(* Logix 5000 project; controller PLC_MCC1300_75F1 vendor 1 type 14 code 166 rev 32.11; software revision 32.04 *)

TASK _18_STI (periodic, rate 10 ms, priority 10, watchdog 500 ms) : _18_STI
TASK Diagnostic (periodic, rate 500 ms, priority 15, watchdog 2000 ms) : Modules
TASK MainTask (periodic, rate 6 ms, priority 10, watchdog 500 ms) : Initialize, MainProgram, CommandLogic, MotionLogic, Communication

MODULES
   Local : vendor 1 type 14 code 166 (ICP 0, rev 32.11)
      ETH_MCC1300 : 1756-EN2T (ICP 1, Ethernet 138.84.12.118, rev 11.1)
         ETH_M2 : 1756-EN2T (Ethernet 138.84.12.123, rev 10.7)   // Plant Network
             : 1756-IB16 (ICP 2, rev 3.4, Input RPI 20 ms)
             : 1756-IB16 (ICP 6, rev 3.4, Input RPI 20 ms)
             : 1756-IB16 (ICP 3, rev 3.4, Input RPI 20 ms)
             : 1756-IB16 (ICP 4, rev 3.4, Input RPI 20 ms)
             : 1756-IB16 (ICP 5, rev 3.4, Input RPI 20 ms)
             : vendor 1 type 7 code 16 (ICP 11, rev 3.4, Output RPI 20 ms)
                 ETH_M2:11:O.Data   // Local output updates
            Rio_Loops_2_3 : 1756-DHRIO (ICP 13, rev 7.2, Input RPI 25 ms)
               VMCC_TD : 1771-ASB (RIO 8, rev 1.1, Output RPI 48 ms)
                    VMCC_TD:O   // RACK 2 OUTPUT UPDATES
               VMCC_M2CM01_SPEED : vendor 1 type 12 code 51 (RIO 13, rev 1.1, Output RPI 48 ms)
                    VMCC_M2CM01_SPEED:O   // RACK 3 OUPUT UPDATES
               VMCC_M2_M2CM02_Speed : vendor 1 type 12 code 51 (RIO 14, rev 1.1, Output RPI 48 ms)
                    VMCC_M2_M2CM02_Speed:O   // RACK 3 OUPUT UPDATES
               ROCKWELL_CAPPING_SYSTEM : vendor 1 type 12 code 51 (RIO 12, rev 1.1, Output RPI 48 ms)
                    ROCKWELL_CAPPING_SYSTEM:O   // RACK 3 OUPUT UPDATES
               PANEL_KD_CS1N : vendor 1 type 12 code 51 (RIO 16, rev 1.1, Output RPI 48 ms)
                    PANEL_KD_CS1N:O   // RACK 11 OUPUT UPDATES
               VMCC_M2_M2CM03_Speed : vendor 1 type 12 code 51 (RIO 15, rev 1.1, Output RPI 48 ms)
                    VMCC_M2_M2CM03_Speed:O   // RACK 3 OUPUT UPDATES
               PANEL_TD_CS1N : 1794-ASB (RIO 18, rev 1.1, Output RPI 48 ms)   // Trim knocker 1
                    PANEL_TD_CS1N:O   // RACK 4 OUPUT UPDATES
               Panel_TS_CS2N : vendor 1 type 12 code 51 (RIO 20, rev 1.1, Output RPI 48 ms)
                    Panel_TS_CS2N:O   // RACK 5 OUPUT UPDATES
               PANEL_TD_CS3N : vendor 1 type 12 code 51 (RIO 22, rev 1.1, Output RPI 48 ms)
                    PANEL_TD_CS3N:O   // RACK 5 OUPUT UPDATES
               PANEL_TD_CS4N : vendor 1 type 12 code 51 (RIO 24, rev 1.1, Output RPI 48 ms)
                    PANEL_TD_CS4N:O   // RACK 6 OUPUT UPDATES
               PANEL_TD_CS5N : vendor 1 type 12 code 51 (RIO 26, rev 1.1, Output RPI 48 ms)
                    PANEL_TD_CS5N:O   // RACK 6 OUPUT UPDATES
               PANEL_TD_CS5S : vendor 1 type 12 code 51 (RIO 28, rev 1.1, Output RPI 48 ms)
                    PANEL_TD_CS5S:I.Data[0].15   // Panel-TD-CS5S Relicance Handoff Sensor (Redundant Sensor on South Side)
                    PANEL_TD_CS5S:O   // RACK 7 OUPUT UPDATES
               PANEL_TD_CS4S : vendor 1 type 12 code 51 (RIO 30, rev 1.1, Output RPI 48 ms)
                    PANEL_TD_CS4S:O   // RACK 7 OUPUT UPDATES
               PANEL_TD_CS3S : vendor 1 type 12 code 51 (RIO 32, rev 1.1, Output RPI 48 ms)
                    PANEL_TD_CS3S:O   // RACK 10 OUPUT UPDATES
               PANEL_TD_CS2S : vendor 1 type 12 code 51 (RIO 34, rev 1.1, Output RPI 48 ms)
                    PANEL_TD_CS2S:O   // RACK 10 OUPUT UPDATES
               BENCHBOARD : vendor 1 type 12 code 51 (RIO 36, rev 1.1, Output RPI 48 ms)
                    BENCHBOARD:O   // RACK 11 OUPUT UPDATES
               PANEL_KD_CS1S : vendor 1 type 12 code 51 (RIO 38, rev 1.1, Output RPI 48 ms)
               PANEL_TD_CS1S : vendor 1 type 12 code 51 (RIO 40, rev 1.1, Output RPI 48 ms)
                    PANEL_TD_CS1S:O   // RACK 12 OUPUT UPDATES
               VMCC_M2CM4S : vendor 1 type 12 code 51 (RIO 42, rev 1.1, Output RPI 48 ms)
                    VMCC_M2CM4S:O   // RACK 12 OUPUT UPDATES
               VMCC_M2_M2CM4N : vendor 1 type 12 code 51 (RIO 43, rev 1.1, Output RPI 48 ms)
                    VMCC_M2_M2CM4N:O   // RACK 12 OUPUT UPDATES
               VMCC_M2_M2CM9S : vendor 1 type 12 code 51 (RIO 52, rev 1.1, Output RPI 48 ms)
                    VMCC_M2_M2CM9S:O   // RACK 15 OUPUT UPDATES
               VMCC_M2_M2CM9N : vendor 1 type 12 code 51 (RIO 53, rev 1.1, Output RPI 48 ms)
                    VMCC_M2_M2CM9N:O   // RACK 15 OUPUT UPDATES
               VMCC_M2_M2CM10S : vendor 1 type 12 code 51 (RIO 54, rev 1.1, Output RPI 48 ms)
                    VMCC_M2_M2CM10S:O   // RACK 15 OUPUT UPDATES
               VMCC_M2_M2CM10N : vendor 1 type 12 code 51 (RIO 55, rev 1.1, Output RPI 48 ms)
                    VMCC_M2_M2CM10N:O   // RACK 15 OUPUT UPDATES
               VMCC_M2_M2CM11S : vendor 1 type 12 code 51 (RIO 56, rev 1.1, Output RPI 48 ms)
                    VMCC_M2_M2CM11S:O   // RACK 16 OUPUT UPDATES
               VMCC_M2_M2CM11N : vendor 1 type 12 code 51 (RIO 57, rev 1.1, Output RPI 48 ms)
                    VMCC_M2_M2CM11N:O   // RACK 16 OUPUT UPDATES
               VMCC_M2_M2CM12S : vendor 1 type 12 code 51 (RIO 58, rev 1.1, Output RPI 48 ms)
                    VMCC_M2_M2CM12S:O   // RACK 16 OUPUT UPDATES
               VMCC_M2_M2CM12N : vendor 1 type 12 code 51 (RIO 59, rev 1.1, Output RPI 48 ms)
                    VMCC_M2_M2CM12N:O   // RACK 16 OUPUT UPDATES
               MB : vendor 1 type 12 code 51 (RIO 60, rev 1.1, Output RPI 48 ms)
                    MB:O   // RACK 17 OUPUT UPDATES
               VMCC_M2_M2CM5S : vendor 1 type 12 code 51 (RIO 44, rev 1.1, Output RPI 48 ms)
                    VMCC_M2_M2CM5S:O   // RACK 13 OUPUT UPDATES
               VMCC_M2_M2CM5N : vendor 1 type 12 code 51 (RIO 45, rev 1.1, Output RPI 48 ms)
                    VMCC_M2_M2CM5N:O   // RACK 13 OUPUT UPDATES
               VMCC_M2_M2CM6S : vendor 1 type 12 code 51 (RIO 46, rev 1.1, Output RPI 48 ms)
                    VMCC_M2_M2CM6S:O   // RACK 13 OUPUT UPDATES
               VMCC_M2_M2CM6N : vendor 1 type 12 code 51 (RIO 47, rev 1.1, Output RPI 48 ms)
                    VMCC_M2_M2CM6N:O   // RACK 13 OUPUT UPDATES
               VMCC_M2_M2CM7S : vendor 1 type 12 code 51 (RIO 48, rev 1.1, Output RPI 48 ms)
                    VMCC_M2_M2CM7S:O   // RACK 14 OUPUT UPDATES
               VMCC_M2_M2CM7N : vendor 1 type 12 code 51 (RIO 49, rev 1.1, Output RPI 48 ms)
                    VMCC_M2_M2CM7N:O   // RACK 14 OUPUT UPDATES
               VMCC_M2_M2CM8S : vendor 1 type 12 code 51 (RIO 50, rev 1.1, Output RPI 48 ms)
                    VMCC_M2_M2CM8S:O   // RACK 14 OUPUT UPDATES
               VMCC_M2_M2CM8N : vendor 1 type 12 code 51 (RIO 51, rev 1.1, Output RPI 48 ms)
                    VMCC_M2_M2CM8N:O   // RACK 14 OUPUT UPDATES
      RIOM13 : 1794-AENTR (Ethernet 192.168.36.11, rev 1.1, Output RPI 20 ms)
         R03_S00 : 1794-IB16 (Flex 0, rev 1.1)
         R03_S01 : 1794-IB16 (Flex 1, rev 1.1)
         R03_S02 : vendor 1 type 7 code 35 (Flex 2, rev 1.1)
      E73AZ1 : vendor 1 type 37 code 49 (Ethernet 192.168.32.131, rev 7.1, MotionDiagnostics RPI 1 ms, MotionSync RPI 1 ms)
      E93AZ1 : vendor 1 type 37 code 49 (Ethernet 192.168.32.132, rev 7.1, MotionDiagnostics RPI 1 ms)
      E53AZ1 : vendor 1 type 45 code 15 (Ethernet 192.168.32.101, rev 2.3, AMotionDiagnostics RPI 1 ms)
      E61AZ1 : vendor 1 type 45 code 15 (Ethernet 192.168.32.102, rev 2.3, AMotionDiagnostics RPI 1 ms)
      E62AZ1 : vendor 1 type 45 code 15 (Ethernet 192.168.32.103, rev 2.3, AMotionDiagnostics RPI 1 ms)
      E63AZ1 : vendor 1 type 45 code 15 (Ethernet 192.168.32.104, rev 2.3, AMotionDiagnostics RPI 1 ms)
      E64AZ1 : vendor 1 type 45 code 15 (Ethernet 192.168.32.105, rev 2.3, AMotionDiagnostics RPI 1 ms)
      E65AZ1 : vendor 1 type 45 code 15 (Ethernet 192.168.32.106, rev 2.3, AMotionDiagnostics RPI 1 ms)
      E66AZ1 : vendor 1 type 45 code 15 (Ethernet 192.168.32.107, rev 2.3, AMotionDiagnostics RPI 1 ms)
      E67AZ1 : vendor 1 type 45 code 15 (Ethernet 192.168.32.108, rev 2.3, AMotionDiagnostics RPI 1 ms)
      E71AZ1 : vendor 1 type 45 code 15 (Ethernet 192.168.32.109, rev 2.3, AMotionDiagnostics RPI 1 ms)
      E76AZ1 : vendor 1 type 45 code 15 (Ethernet 192.168.32.110, rev 2.3, AMotionDiagnostics RPI 1 ms)
      E77AZ1 : vendor 1 type 45 code 15 (Ethernet 192.168.32.111, rev 2.3, AMotionDiagnostics RPI 1 ms)
      E78AZ1 : vendor 1 type 45 code 15 (Ethernet 192.168.32.112, rev 2.3, AMotionDiagnostics RPI 1 ms)
      E81AZ1 : vendor 1 type 45 code 15 (Ethernet 192.168.32.113, rev 2.3, AMotionDiagnostics RPI 1 ms)
      E82AZ1 : vendor 1 type 45 code 15 (Ethernet 192.168.32.114, rev 2.3, AMotionDiagnostics RPI 1 ms)
      E83AZ1 : vendor 1 type 45 code 15 (Ethernet 192.168.32.115, rev 2.3, AMotionDiagnostics RPI 1 ms)
      E84AZ1 : vendor 1 type 45 code 15 (Ethernet 192.168.32.116, rev 2.3, AMotionDiagnostics RPI 1 ms)
      E85AZ1 : vendor 1 type 45 code 15 (Ethernet 192.168.32.117, rev 2.3, AMotionDiagnostics RPI 1 ms)
      E86AZ1 : vendor 1 type 45 code 15 (Ethernet 192.168.32.118, rev 2.3, AMotionDiagnostics RPI 1 ms)
      E87AZ1 : vendor 1 type 45 code 15 (Ethernet 192.168.32.119, rev 2.3, AMotionDiagnostics RPI 1 ms)
      E88AZ1 : vendor 1 type 45 code 15 (Ethernet 192.168.32.120, rev 2.3, AMotionDiagnostics RPI 1 ms)
      E91AZ1 : vendor 1 type 45 code 15 (Ethernet 192.168.32.121, rev 2.3, AMotionDiagnostics RPI 1 ms)
      E96AZ1 : vendor 1 type 45 code 15 (Ethernet 192.168.32.122, rev 2.3, AMotionDiagnostics RPI 1 ms)
      E97AZ1 : vendor 1 type 45 code 15 (Ethernet 192.168.32.123, rev 2.3, AMotionDiagnostics RPI 1 ms)
      E98AZ1 : vendor 1 type 45 code 15 (Ethernet 192.168.32.124, rev 2.3, AMotionDiagnostics RPI 1 ms)
      M3AZ01 : vendor 1 type 45 code 15 (Ethernet 192.168.32.141, rev 2.3, AMotionDiagnostics RPI 1 ms)
      M3AZ02 : vendor 1 type 45 code 15 (Ethernet 192.168.32.142, rev 2.3, AMotionDiagnostics RPI 1 ms)
      M3AZ03 : vendor 1 type 45 code 15 (Ethernet 192.168.32.143, rev 2.3, AMotionDiagnostics RPI 1 ms)
      M3AZ04 : vendor 1 type 45 code 15 (Ethernet 192.168.32.144, rev 2.3, AMotionDiagnostics RPI 1 ms)
      M3AZ05 : vendor 1 type 45 code 15 (Ethernet 192.168.32.145, rev 2.3, AMotionDiagnostics RPI 1 ms)
      M3AZ06 : vendor 1 type 45 code 15 (Ethernet 192.168.32.146, rev 2.3, AMotionDiagnostics RPI 1 ms)
      M3AZ07 : vendor 1 type 45 code 15 (Ethernet 192.168.32.147, rev 2.3, AMotionDiagnostics RPI 1 ms)
      M3AZ08 : vendor 1 type 45 code 15 (Ethernet 192.168.32.148, rev 2.3, AMotionDiagnostics RPI 1 ms)
      M3AZ09 : vendor 1 type 45 code 15 (Ethernet 192.168.32.149, rev 2.3, AMotionDiagnostics RPI 1 ms)
      M3AZ10 : vendor 1 type 45 code 15 (Ethernet 192.168.32.150, rev 2.3, AMotionDiagnostics RPI 1 ms)
      D010M1PM1 : vendor 1 type 45 code 15 (Ethernet 192.168.36.131, rev 2.3, AMotionDiagnostics RPI 1 ms)
      D010M2PM1 : vendor 1 type 45 code 15 (Ethernet 192.168.36.132, rev 2.3, AMotionDiagnostics RPI 1 ms)
      D020M1PM1 : vendor 1 type 45 code 15 (Ethernet 192.168.36.133, rev 2.3, AMotionDiagnostics RPI 1 ms)
      TDKAZ00N : vendor 1 type 45 code 15 (Ethernet 192.168.31.101, rev 2.3, AMotionDiagnostics RPI 1 ms)
      TDKAZ00S : vendor 1 type 45 code 15 (Ethernet 192.168.31.102, rev 2.3, AMotionDiagnostics RPI 1 ms)
      TDKAZ01N : vendor 1 type 45 code 15 (Ethernet 192.168.31.103, rev 2.3, AMotionDiagnostics RPI 1 ms)
      TDKAZ01S : vendor 1 type 45 code 15 (Ethernet 192.168.31.104, rev 2.3, AMotionDiagnostics RPI 1 ms)
      TDKAZ02N : vendor 1 type 45 code 15 (Ethernet 192.168.31.105, rev 2.3, AMotionDiagnostics RPI 1 ms)
      TDKAZ02S : vendor 1 type 45 code 15 (Ethernet 192.168.31.106, rev 2.3, AMotionDiagnostics RPI 1 ms)
      TDKAZ03N : vendor 1 type 45 code 15 (Ethernet 192.168.31.107, rev 2.3, AMotionDiagnostics RPI 1 ms)
      TDKAZ03S : vendor 1 type 45 code 15 (Ethernet 192.168.31.108, rev 2.3, AMotionDiagnostics RPI 1 ms)
      TDKAZ04N : vendor 1 type 45 code 15 (Ethernet 192.168.31.109, rev 2.3, AMotionDiagnostics RPI 1 ms)
      TDKAZ04S : vendor 1 type 45 code 15 (Ethernet 192.168.31.110, rev 2.3, AMotionDiagnostics RPI 1 ms)
      TDKAZ05N : vendor 1 type 45 code 15 (Ethernet 192.168.31.111, rev 2.3, AMotionDiagnostics RPI 1 ms)
      TDKAZ05S : vendor 1 type 45 code 15 (Ethernet 192.168.31.112, rev 2.3, AMotionDiagnostics RPI 1 ms)
      TDAZ00N : vendor 1 type 45 code 15 (Ethernet 192.168.31.113, rev 2.3, AMotionDiagnostics RPI 1 ms)
      TDAZ00S : vendor 1 type 45 code 15 (Ethernet 192.168.31.114, rev 2.3, AMotionDiagnostics RPI 1 ms)
      TDAZ01N : vendor 1 type 45 code 15 (Ethernet 192.168.31.115, rev 2.3, AMotionDiagnostics RPI 1 ms)
      TDAZ01S : vendor 1 type 45 code 15 (Ethernet 192.168.31.116, rev 2.3, AMotionDiagnostics RPI 1 ms)
      TDAZ02N : vendor 1 type 45 code 15 (Ethernet 192.168.31.117, rev 2.3, AMotionDiagnostics RPI 1 ms)
      TDAZ02S : vendor 1 type 45 code 15 (Ethernet 192.168.31.118, rev 2.3, AMotionDiagnostics RPI 1 ms)
      TDAZ03N : vendor 1 type 45 code 15 (Ethernet 192.168.31.119, rev 2.3, AMotionDiagnostics RPI 1 ms)
      TDAZ03S : vendor 1 type 45 code 15 (Ethernet 192.168.31.120, rev 2.3, AMotionDiagnostics RPI 1 ms)
      TDAZ04N : vendor 1 type 45 code 15 (Ethernet 192.168.31.121, rev 2.3, AMotionDiagnostics RPI 1 ms)
      TDAZ04S : vendor 1 type 45 code 15 (Ethernet 192.168.31.122, rev 2.3, AMotionDiagnostics RPI 1 ms)
      TDAZ05N : vendor 1 type 45 code 15 (Ethernet 192.168.31.123, rev 2.3, AMotionDiagnostics RPI 1 ms)
      TDAZ05S : vendor 1 type 45 code 15 (Ethernet 192.168.31.124, rev 2.3, AMotionDiagnostics RPI 1 ms)
      E152AP1 : vendor 1 type 12 code 317 (Ethernet 192.168.32.11, rev 4.1)
         R00_S03 : 5069-IB16 (5069 3, rev 2.1, StandardDataDriven RPI 5 ms)
         R00_S04 : 5069-IB16 (5069 4, rev 2.1, StandardDataDriven RPI 5 ms)
         R00_S02 : 5069-IB16 (5069 2, rev 2.1, StandardDataDriven RPI 5 ms)
         R00_S01 : 5069-IB16 (5069 1, rev 2.1, StandardDataDriven RPI 5 ms)
         R00_S05 : 5069-IB16 (5069 5, rev 2.1, StandardDataDriven RPI 5 ms)
         R00_S06 : 5069-IB16 (5069 6, rev 2.1, StandardDataDriven RPI 5 ms)
         R00_S07 : 5069-IB16 (5069 7, rev 2.1, StandardDataDriven RPI 5 ms)
         R00_S08 : 5069-IB16 (5069 8, rev 2.1, StandardDataDriven RPI 5 ms)
         R00_S09 : 5069-IB16 (5069 9, rev 2.1, StandardDataDriven RPI 5 ms)
         R00_S10 : 5069-IB16 (5069 10, rev 2.1, StandardDataDriven RPI 5 ms)
         R00_S11 : 5069-IB16 (5069 11, rev 2.1, StandardDataDriven RPI 5 ms)
         R00_S12 : 5069-IB16 (5069 12, rev 2.1, StandardDataDriven RPI 5 ms)
         R00_S13 : 5069-OB16 (5069 13, rev 3.1, StandardDataDriven RPI 5 ms)
         R00_S14 : 5069-OB16 (5069 14, rev 3.1, StandardDataDriven RPI 5 ms)
         R00_S15 : 5069-OB16 (5069 15, rev 3.1, StandardDataDriven RPI 5 ms)
         R00_S16 : 5069-OB16 (5069 16, rev 3.1, StandardDataDriven RPI 5 ms)
         R00_S17 : 5069-OB16 (5069 17, rev 3.1, StandardDataDriven RPI 5 ms)
      M3683AP1 : vendor 1 type 12 code 317 (Ethernet 192.168.31.12, rev 4.1)
         R01_S01 : 5069-IB16 (5069 1, rev 2.1, StandardDataDriven RPI 5 ms)
         R01_S02 : 5069-IB16 (5069 2, rev 2.1, StandardDataDriven RPI 5 ms)
         R01_S03 : 5069-IB16 (5069 3, rev 2.1, StandardDataDriven RPI 5 ms)
         R01_S04 : 5069-IB16 (5069 4, rev 2.1, StandardDataDriven RPI 5 ms)
         R01_S05 : 5069-OB16 (5069 5, rev 3.1, StandardDataDriven RPI 5 ms)
         R01_S06 : 5069-OB16 (5069 6, rev 3.1, StandardDataDriven RPI 5 ms)
         R01_S07 : 5069-OB16 (5069 7, rev 3.1, StandardDataDriven RPI 5 ms)
         R01_S08 : 5069-OB16 (5069 8, rev 3.1, StandardDataDriven RPI 5 ms)
         R01_S09 : 5069-OB16 (5069 9, rev 3.1, StandardDataDriven RPI 5 ms)
         R01_S10 : 5069-IB16 (5069 10, rev 2.1, StandardDataDriven RPI 5 ms)
      TD5680AP1 : vendor 1 type 12 code 317 (Ethernet 192.168.31.11, rev 4.1)
         R02_S01 : 5069-IB16 (5069 1, rev 2.1, StandardDataDriven RPI 5 ms)
         R02_S02 : 5069-IB16 (5069 2, rev 2.1, StandardDataDriven RPI 5 ms)
         R02_S03 : 5069-OB16 (5069 3, rev 3.1, StandardDataDriven RPI 5 ms)
         R02_S04 : 5069-OB16 (5069 4, rev 3.1, StandardDataDriven RPI 5 ms)
         R02_S05 : 5069-OB16 (5069 5, rev 3.1, StandardDataDriven RPI 5 ms)
         R02_S06 : 5069-OB16 (5069 6, rev 3.1, StandardDataDriven RPI 5 ms)
         R02_S07 : 5069-IB16 (5069 7, rev 2.1, StandardDataDriven RPI 5 ms)
         R02_S08 : 5069-IB16 (5069 8, rev 2.1, StandardDataDriven RPI 5 ms)
END_MODULES

TYPE AUX_COSTANTS :
STRUCT
   dM302SnapOffset_cmm : DINT;   // Distance from origin sepoint and snapbar [mm/100]
   dM302SpeedUpMinGapInConvoy_cmm : DINT;   // Minimum gap in convoy [mm/100]
   dM310_PopUpCycleTime_s : DINT[2];   // Popup cycle time [s]
   dM315_PopUpCycleTime_s : DINT[2];   // Popup cycle time [s]
END_STRUCT
END_TYPE

TYPE CM_AreaStackerToLine :
STRUCT
   dSyncHead : DINT;
   xRequestAccessArea : BOOL;
   xAccessAreaAccepted : BOOL;
   xAreaOk : BOOL;
   xStackerInUnloaderMode : BOOL;
   xStackerInProduction : BOOL;
   xPlateOnFrame : BOOL[32];
   xSB_SilenceAlarm : BOOL;
   xSB_SendToCullet : BOOL;
   xSB_LineCycle : BOOL;
   xSB_StopLineCycle : BOOL;
   xSB_LineJogPlus : BOOL;
   xSB_LineJogMinus : BOOL;
   xSB_DestinationChange : BOOL;
   iPresetNumberPlateOnRack : INT[2];
   iActualNumberPlateOnRack : INT[2];
   iPresetNumberPlateAddOnRack : INT[2];
   iActualNumberPlateAddOnRack : INT[2];
   dGap_cmm : DINT;
   dMsgDataSyncFdbk : DINT;
   dMsgDataSync : DINT;
   dMsgOPTSyncFdbk : DINT;
   dMsgOPTSync : DINT;
   dSyncTail : DINT;
END_STRUCT
END_TYPE

TYPE CM_ConveyorStackerToLine :
STRUCT
   dSyncHead : DINT;
   xCycleOn : BOOL;
   xConditionOkForStopCycle : BOOL;
   xInitialContionOk : BOOL;
   xOutputEnable : BOOL;
   xReadyToMove : BOOL;
   xFeedbackRotation : BOOL;
   xRequestReturnInLine : BOOL;
   xRequestUnload : BOOL;
   xRotationForUnload : BOOL;
   xRotationForLoad : BOOL;
   xEndPhaseLoad : BOOL;
   xManualCommandFwd : BOOL;
   xManualCommandBkw : BOOL;
   xAirMode : BOOL;
   xTinMode : BOOL;
   xPhotocell1 : BOOL;
   xPhotocell2 : BOOL;
   xPlateOnConveyor : BOOL[32];
   dSyncTail : DINT;
END_STRUCT
END_TYPE

TYPE CM_DATA_Z200 :   // Cap data coming from Z200
STRUCT
   dSyncHead : DINT;   // Synchro head
   tConvoyCap : UDT_ConvoyCap_ZC;   // Cap data
   dSyncTail : DINT;   // Synchro tail
END_STRUCT
END_TYPE

TYPE CM_INPUT_Z200 :
STRUCT
   dSyncHead : DINT;   // Synchro head
   xZ200_CycleON : BOOL;   // Z200 Cycle ON
   xSnapDone : BOOL;   // Snap done
   xSBStartEmptyingZ301 : BOOL;   // CS4201 Start Emptying Z301 Button
   xSBStopEmptyingZ301 : BOOL;   // CS4201 Stop Emptying Z301 Button
   xSBResetAnomalyZ301 : BOOL;   // CS4201 Reset Anomaly Z301 Button
   xResetGeneralEmergency : BOOL;   // Reset General Emergency
   xCrossbreakActive : BOOL;   // Crossbreak Active
   xEmergencyON : BOOL;   // Emergency ON
   xMainCulletConveyorAllow : BOOL;   // Main Cullet Conveyor Allow
   dLehrSpeed_mm_min : DINT;   // Lehr speed [mm/min]
   dDataSync : DINT;   // Snap cap data sent
   rgdSpare : DINT[10];
   dSyncTail : DINT;   // Synchro tail
END_STRUCT
END_TYPE

TYPE CM_LineToAreaStacker :
STRUCT
   dSyncHead : DINT;
   xConditionOkForAccessArea : BOOL;
   xSBSendToCullet : BOOL;
   xSBLineCycle : BOOL;
   xSBStopLineCycle : BOOL;
   xHLAlarmStartLineCycle : BOOL;
   xSBChangeDestination : BOOL;
   dMsgDataSyncFdbk : DINT;
   dMsgDataSync : DINT;
   dMsgOPTSyncFdbk : DINT;
   dMsgOPTSync : DINT;
   dSyncTail : DINT;
END_STRUCT
END_TYPE

TYPE CM_LineToConveyorStacker :
STRUCT
   dSyncHead : DINT;
   xEmergencyOn : BOOL;
   xLineCycleOn : BOOL;
   xLineStopCycle : BOOL;
   xRequestForceStop : BOOL;
   xResetAlarms : BOOL;
   xResetEmergency : BOOL;
   xPowerOnByLine : BOOL;
   xInitialConditionOk : BOOL;
   xOutputEnable : BOOL;
   xReadyToMove : BOOL;
   xFeedbackRotation : BOOL;
   xEndPhaseLoad : BOOL;
   xRotationForLoad : BOOL;
   xRequestForUnload : BOOL;
   xRotationForUnload : BOOL;
   xManualCommandFwd : BOOL;
   xManualCommandBkw : BOOL;
   xSendToCullet : BOOL;
   xLineJogPlus : BOOL;
   xLineJogMinus : BOOL;
   dLineSpeed_dmm_min : DINT;
   dSyncTail : DINT;
END_STRUCT
END_TYPE

TYPE CM_OUTPUT_Z200 :
STRUCT
   dSyncHead : DINT;   // Synchro head
   xZ300_CycleON : BOOL;   // Z300 Cycle ON
   xBLStartEmptyingZ301Light : BOOL;   // CS4201 Start Emptying Z301 Button Light
   xBLStopEmptyingZ301Light : BOOL;   // CS4201 Stop Emptying Z301 Button Light
   xBLAnomalyZ301Light : BOOL;   // CS4201 Anomaly Z301 Button Light
   xBLAnomalyZ302Light : BOOL;   // CS4201 Anomaly Z302 Button Light
   dDataSyncFdbk : DINT;   // Snap cap sync feedback
   dLineSpeed_mm_min : DINT;   // Line speed [mm/min]
   rgdSpare : DINT[10];
   dSyncTail : DINT;   // Synchro tail
END_STRUCT
END_TYPE

TYPE DATA_CAP_PILKINGTON :
STRUCT
   dHost_ID : DINT;   // Host ID
   dCap_Length_64ths : DINT;   // Cap Length (64ths)
   dCap_Primary_Destination_Mask : DINT;   // Cap Primary Destination Mask
   Packing_station_1_Mask : DINT;   // Packing Station 1 Mask
   Packing_station_2_Mask : DINT;   // Packing Station 2 Mask
   Packing_station_3_Mask : DINT;   // Packing Station 3 Mask
   Packing_station_4_Mask : DINT;   // Packing Station 4 Mask
   Packing_station_5_Mask : DINT;   // Packing Station 5 Mask
   dSplit_A_Width_64ths : DINT;   // Split A Width (64ths)
   dSplit_A_Dest_Mask : DINT;   // Split A Destination Mask
   dSplit_B_Width_64ths : DINT;   // Split B Width (64ths)
   dSplit_B_Dest_Mask : DINT;   // Split B Destination Mask
   dSplit_C_Width_64ths : DINT;   // Split C Width (64ths)
   dSplit_C_Dest_Mask : DINT;   // Split C Destination Mask
   dSplit_D_Width_64ths : DINT;   // Split D Width (64ths)
   dSplit_D_Dest_Mask : DINT;   // Split D Destination Mask
   dCap_Secondary_Dest_Mask : DINT;   // Cap Secondary Destination Mask
   dTrim_Home_Side_64ths : DINT;   // Trim on home (left) side (64ths)
   dTrim_Far_Side_64ths : DINT;   // Trim on far (right) side (64ths)
   dControl_Bits_For_Legs : DINT;   // Control bits for legs
   dCap_Width_64ths : DINT;   // Cap Width (64ths)
   dReject_Mask : DINT;   // Split Reject mask
   dPattern_number : DINT;   // Pattern number
   dSpare1 : DINT;   // Spare
   dSpare2 : DINT;   // Spare
   dSpare3 : DINT;   // Spare
   dMainline_History_Word : DINT;   // Mainline History Word
   dSpare4 : DINT;   // Spare
   dSpare5 : DINT;   // Spare
   dSpare6 : DINT;   // Spare
   dSpare7 : DINT;   // Spare
   dSpare8 : DINT;   // Spare
   dSpare9 : DINT;   // Spare
END_STRUCT
END_TYPE

TYPE GP_AccessArea_STC :
STRUCT
   ST_xAccessRequest : BOOL;
   ST_xAccessAccepted : BOOL;
   ST_xAccessAnnulled : BOOL;
   ST_xAccessAcceptedAndButtonReleased : BOOL;
   ST_xConditionOkForAccess : BOOL;
   ST_xDelayForceAccess : BOOL;
   ST_xSafetyOkForCycle : BOOL;
   OSR_xAccessRequest : BOOL;
   OSR_xAccessAcceptedAndButtonReleased : BOOL;
   OSR_xRemoveAccess : BOOL;
   OSR_xRemoveAccessNotAccepted : BOOL;
   OS_xAccessRequest : BOOL;
   OS_xSafetyOK : BOOL;
   tmON_ForceAccess : TIMER;
END_STRUCT
END_TYPE

TYPE GP_NetworkDiag_v1 :
STRUCT
   sModuleName : STRING;   // Module name
   xConnected : BOOL;   // Module connected
   xFaulted : BOOL;   // Module faulted
   dEntryStatus : DINT;
   dFaultCode : DINT;
   dFaultInfo : DINT;
   dInstance : DINT;
END_STRUCT
END_TYPE

TYPE GP_OB_Initialize_STC :
STRUCT
   dElapsed_1h_ms : DINT;   // Decimal
   dElapsed_1min_ms : DINT;   // Decimal
   dElapsed_1s_ms : DINT;   // Decimal
   dElapsed_2min_ms : DINT;   // Decimal
   dElapsed_2s_ms : DINT;   // Decimal
   dElapsed_5s_ms : DINT;   // Decimal
   dElapsed_10min_ms : DINT;   // Decimal
   dElapsed_10s_ms : DINT;   // Decimal
   dElapsed_30min_ms : DINT;   // Decimal
   dElapsed_30s_ms : DINT;   // Decimal
   dElapsed_100ms_ms : DINT;   // Decimal
   dElapsed_200ms_ms : DINT;   // Decimal
   dElapsed_400ms_ms : DINT;   // Decimal
   dElapsed_500ms_ms : DINT;   // Decimal
   dElapsed_800ms_ms : DINT;   // Decimal
   dlLastExecValue_us : DINT;   // Decimal
   rReminder_ms : REAL;   // Float
   lwOldStartTime : DINT[2];   // Old start time execution
   lwStartTime : DINT[2];   // Start time execution
END_STRUCT
END_TYPE

TYPE GP_TrackingSearchPlate_STC :
STRUCT
   rgdHeadPointer : DINT[5];   // Head pointer
   rgdTailPointer : DINT[5];   // Tail pointer
   rgdHead_cmm : DINT[5];   // Head position [cmm]
   rgdTail_cmm : DINT[5];   // Tail position [cmm]
   rgxHead : DINT;   // Head found
   rgxTail : DINT;   // Tail found
   xHeadPresence : BOOL;   // At least one head
   xTailPresence : BOOL;   // At least one tail
END_STRUCT
END_TYPE

TYPE HMI_LiteData :
STRUCT
   dHead_PosX_mm : DINT;   // Plate head position X [mm]
   dTail_PosX_mm : DINT;   // Plate tail position X [mm]
   dPlateLength_mm : DINT;   // Plate length [mm]
   dPositionY_mm : DINT;   // Plate position Y [mm]- Operator side
   dPlateWidth_mm : DINT;   // Plate widht [mm]
   dPlateId : DINT;   // Plate ID
   dProductionID : DINT;   // Production ID
   dSource : DINT;   // Plate source
   dDestination : DINT;   // Plate Main destination
   dAlternative : DINT;   // Plate Alternative destination
   dSecondDestination : DINT;   // Plate 2nd choice destination
END_STRUCT
END_TYPE

TYPE MAC_Conveyor :
STRUCT
   ST_xInitialConditionOK : BOOL;   // Initial condition OK
   ST_xInitialConditionOK_BW : BOOL;   // Initial condition OK backward
   ST_xCleaningConditionOK : BOOL;   // Cleaning condition OK
   ST_xCleaningAccepted : BOOL;   // Cleaning accepted
   ST_xReqCleaning : BOOL;   // Request cleaning
   ST_xPlatePresence : BOOL;   // Plate presence memory
   ST_xPhasesInProgress : BOOL;   // Phases in progress
   ST_xCycleLoadUnload : BOOL;   // Cycle load/unload simultaneously
   ST_xStopMachineFault : BOOL;   // Stopped machine fault
   ST_xStopNextCycleFault : BOOL;   // Stop next cycle fault
   ST_xConditionOKStopCycle : BOOL;   // Condition OK for stop cycle
   ST_xOutputEnable : BOOL;   // Output enable
   ST_xMachineAlarm : BOOL;   // Machine alarm
   ST_xMachineWarning : BOOL;   // Machine warning
   ST_xIdPlatePresence : BOOL;   // Id plate presence
   ST_xFeedbackRotation : BOOL;   // Feedback rotation
   ST_xRampInProgress : BOOL;   // Ramp in progress
   ST_xAccInProgress : BOOL;   // Acceleration in progress
   ST_xDecInProgress : BOOL;   // Deceleration in progress
   ST_xWaitStopNextMachine : BOOL;   // Wait stop next machine
   ST_xWaitMachineStop : BOOL;   // Wait machine stop
   ST_xWaitReadyToMove : BOOL;   // Wait ready to move
   ST_xEnableControlError : BOOL;   // Enable control error
   ST_xManualMode : BOOL;   // Manual mode enabled
   ST_xPlateSynchronized : BOOL;   // Plate synchronized
   ST_xVirtualDoorEnabled : BOOL;   // Virtual door enabled
   ST_xDisableLoadUnloadOnStop : BOOL;   // Temporary disable of load/unload continuosly after a bit wait machine stop
   ST_xPlatePassageUpstream_FW : BOOL;   // Plate in passage upstream
   ST_xPlatePassageUpstream_BKW : BOOL;   // Plate in passage upstream
   ST_xPlatePassageDownstream_FW : BOOL;   // Plate in passage downstream
   ST_xPlatePassageDownstream_BKW : BOOL;   // Plate in passage downstream
   ST_xAxleReadyToMoveDelayed : BOOL;   // Axle ready to move delayed (NU)
   ST_xSafetyMovement : BOOL;   // Safety Mouvement
   ST_xReqDescent : BOOL;   // popup conveyor
   ST_xPhaseError : BOOL;   // Phase error, send lites to cullet
   ST_xAux1 : BOOL;   // ST Aux 1
   ST_xAux2 : BOOL;   // ST Aux 2
   ST_xAux3 : BOOL;   // ST Aux 3
   ST_xAux4 : BOOL;   // ST Aux 4
   OSR_xUnload : BOOL;   // OSR Unload
   OSR_xSynchroPhotocellHead : BOOL;   // OSR Synchronization photocell head
   OSR_xSynchroPhotocellTail : BOOL;   // OSR Synchronization photocell tail
   OSR_xPosReq : BOOL;   // OSR Positioning request
   OS_xLoad_FW : BOOL;   // OS Load forward
   OS_xUnload_FW : BOOL;   // OS Unload forward
   OS_xLoad_BW : BOOL;   // OS Load backward
   OS_xUnload_BW : BOOL;   // OS Unload backward
   OS_xUnpack : BOOL;   // OS Unpack convoy
   OS_xSynchroPhotocellHead : BOOL;   // OS Synchronization photocell head
   OS_xSynchroPhotocellTail : BOOL;   // OS Synchronization photocell tail
   OS_xChangeSpeed : BOOL;   // OS Dynamic change speed
   PH_x : DINT;   // Phases
   INPUT_xSyncroPhotocell_1 : BOOL;   // Sincro photocell / start count #1
   INPUT_xSyncroPhotocell_2 : BOOL;   // Sincro photocell / start count #2
   INPUT_xSquaringPhotocell_1 : BOOL;   // Squaring photocell #1
   INPUT_xSquaringPhotocell_2 : BOOL;   // Squaring photocell #2
   INPUT_xSquaringPhotocell_3 : BOOL;   // Squaring photocell #3
   INPUT_xSquaringPhotocell_4 : BOOL;   // Squaring photocell #4
   INPUT_xHighPositionSquaring_1 : BOOL;   // High position squaring #1
   INPUT_xLowPositionSquaring_1 : BOOL;   // Low position squaring #1
   INPUT_xHighPositionSquaring_2 : BOOL;   // High position squaring #2
   INPUT_xLowPositionSquaring_2 : BOOL;   // Low position squaring #2
   INPUT_xHighPositionPopup_1 : BOOL;   // High position pop-up
   INPUT_xLowPositionPopup_1 : BOOL;   // Low position pop-up
   INPUT_xHighPositionPopup_2 : BOOL;   // High position pop-up
   INPUT_xLowPositionPopup_2 : BOOL;   // Low position pop-up
   INPUT_xBrakingResistor_M1 : BOOL;   // Braking resistor
   INPUT_xDriveError_M1 : BOOL;   // Drive error
   INPUT_xDriveFeedback_M1 : BOOL;   // Drive feedback
   INPUT_xDriveInhibit_M1 : BOOL;   // Drive inhibit
   INPUT_xDriveReady_M1 : BOOL;   // Drive ready
   INPUT_xLocalSafetySwitch_M1 : BOOL;   // Local safety switch
   INPUT_xMotorThermalProbe_M1 : BOOL;   // Motor thermal probe
   INPUT_xProtectionMotor_M1 : BOOL;   // Protection motor
   INPUT_xBrakingResistor_M2 : BOOL;   // Braking resistor
   INPUT_xDriveError_M2 : BOOL;   // Drive error
   INPUT_xDriveFeedback_M2 : BOOL;   // Drive feedback
   INPUT_xDriveInhibit_M2 : BOOL;   // Drive inhibit
   INPUT_xDriveReady_M2 : BOOL;   // Drive ready
   INPUT_xLocalSafetySwitch_M2 : BOOL;   // Local safety switch
   INPUT_xMotorThermalProbe_M2 : BOOL;   // Motor thermal probe
   INPUT_xProtectionMotor_M2 : BOOL;   // Protection motor
   INPUT_xBrakingResistor_M3 : BOOL;   // Braking resistor
   INPUT_xDriveError_M3 : BOOL;   // Drive error
   INPUT_xDriveFeedback_M3 : BOOL;   // Drive feedback
   INPUT_xDriveInhibit_M3 : BOOL;   // Drive inhibit
   INPUT_xDriveReady_M3 : BOOL;   // Drive ready
   INPUT_xLocalSafetySwitch_M3 : BOOL;   // Local safety switch
   INPUT_xMotorThermalProbe_M3 : BOOL;   // Motor thermal probe
   INPUT_xProtectionMotor_M3 : BOOL;   // Protection motor
   INPUT_xBrakingResistor_M4 : BOOL;   // Braking resistor
   INPUT_xDriveError_M4 : BOOL;   // Drive error
   INPUT_xDriveFeedback_M4 : BOOL;   // Drive feedback
   INPUT_xDriveInhibit_M4 : BOOL;   // Drive inhibit
   INPUT_xDriveReady_M4 : BOOL;   // Drive ready
   INPUT_xLocalSafetySwitch_M4 : BOOL;   // Local safety switch
   INPUT_xMotorThermalProbe_M4 : BOOL;   // Motor thermal probe
   INPUT_xProtectionMotor_M4 : BOOL;   // Protection motor
   INPUT_xProtectionLiftingFrame_1 : BOOL;   // Protection lifting frame
   INPUT_xFeedBackLiftingFrame_1 : BOOL;   // Feedback lifting frame
   INPUT_xProtectionFan_1 : BOOL;   // Protection fan
   INPUT_xFeedbackVentilation_1 : BOOL;   // Feedback ventilation
   INPUT_xProtectionLiftingFrame_2 : BOOL;   // Protection lifting frame
   INPUT_xFeedBackLiftingFrame_2 : BOOL;   // Feedback lifting frame
   INPUT_xProtectionFan_2 : BOOL;   // Protection fan
   INPUT_xFeedbackVentilation_2 : BOOL;   // Feedback ventilation
   OUTPUT_xRisePopup_1 : BOOL;   // Rise popup #1
   OUTPUT_xDescentPopup_1 : BOOL;   // Descent popup #1
   OUTPUT_xRisePopup_2 : BOOL;   // Rise popup #2
   OUTPUT_xDescentPopup_2 : BOOL;   // Descent popup #2
   OUTPUT_xRiseSquaring_1 : BOOL;   // Rise squaring #1
   OUTPUT_xDescentSquaring_1 : BOOL;   // Descent squaring #1
   OUTPUT_xRiseSquaring_2 : BOOL;   // Rise squaring #2
   OUTPUT_xDescentSquaring_2 : BOOL;   // Descent squaring #2
   OUTPUT_xDriveEnable_M1 : BOOL;   // Drive enable
   OUTPUT_xPositioning_M1 : BOOL;   // Positiong
   OUTPUT_xReverse_M1 : BOOL;   // Reserve
   OUTPUT_xRun_M1 : BOOL;   // Run
   OUTPUT_xDriveEnable_M2 : BOOL;   // Drive enable
   OUTPUT_xPositioning_M2 : BOOL;   // Positiong
   OUTPUT_xReverse_M2 : BOOL;   // Reserve
   OUTPUT_xRun_M2 : BOOL;   // Run
   OUTPUT_xDriveEnable_M3 : BOOL;   // Drive enable
   OUTPUT_xPositioning_M3 : BOOL;   // Positiong
   OUTPUT_xReverse_M3 : BOOL;   // Reserve
   OUTPUT_xRun_M3 : BOOL;   // Run
   OUTPUT_xDriveEnable_M4 : BOOL;   // Drive enable
   OUTPUT_xPositioning_M4 : BOOL;   // Positiong
   OUTPUT_xReverse_M4 : BOOL;   // Reserve
   OUTPUT_xRun_M4 : BOOL;   // Run
   OUTPUT_xFanCommand : BOOL;   // Fan command
   AUX_dPresetStopLoad_cmm : DINT;   // Preset Stop Load position [mm/100]
   AUX_dPresetStopUnload_cmm : DINT;   // Preset Stop Unload position [mm/100]
   AUX_dAccSpace_cmm : DINT;   // Acceleration Space [mm/100]
   AUX_dDecSpace_cmm : DINT;   // Acceleration Space [mm/100]
   AUX_dReqSpeed_mm_min : DINT;   // Conveyor requested speed [mm/min]
   AUX_dAbsPosTarget_M1_cmm : DINT;   // Absolute positioning target [mm/100]
   AUX_dAbsPosTarget_M2_cmm : DINT;   // Absolute positioning target [mm/100]
   AUX_dAbsPosTarget_M3_cmm : DINT;   // Absolute positioning target [mm/100]
   AUX_dAbsPosTarget_M4_cmm : DINT;   // Absolute positioning target [mm/100]
   AUX_dPhPosTarget_cmm : DINT;   // Photocell positioning target [mm/100]
   AUX_dPhPosTarget_2_cmm : DINT;   // Photocell positioning target 2 [mm/100]
   TmON_AxleReadyToMoveDelayed : TIMER;   // Axle ready to move delayed (NU)
   tmON_FeedbackTimeOut_M1 : TIMER;   // Feedback time out
   tmON_DriveInhibit_M1 : TIMER;   // Inhibit time out
   tmOF_DriveEnable_M1 : TIMER;   // Drive enable timer
   tmOF_PowerSaving_M1 : TIMER;   // Power saving timer
   tmON_FeedbackTimeOut_M2 : TIMER;   // Feedback time out
   tmON_DriveInhibit_M2 : TIMER;   // Inhibit time out
   tmOF_DriveEnable_M2 : TIMER;   // Drive enable timer
   tmOF_PowerSaving_M2 : TIMER;   // Power saving timer
   tmON_FeedbackTimeOut_M3 : TIMER;   // Feedback time out
   tmON_DriveInhibit_M3 : TIMER;   // Inhibit time out
   tmOF_DriveEnable_M3 : TIMER;   // Drive enable timer
   tmOF_PowerSaving_M3 : TIMER;   // Power saving timer
   tmON_FeedbackTimeOut_M4 : TIMER;   // Feedback time out
   tmON_DriveInhibit_M4 : TIMER;   // Inhibit time out
   tmOF_DriveEnable_M4 : TIMER;   // Drive enable timer
   tmOF_PowerSaving_M4 : TIMER;   // Power saving timer
   tmON_PosTimeOut_1 : TIMER;   // Positioning timeout 1
   tmON_PosTimeOut_2 : TIMER;   // Positioning timeout 2
   tmON_PosTimeOut_3 : TIMER;   // Positioning timeout 3
   tmON_PosTimeOut_4 : TIMER;   // Positioning timeout 3
   tmON_Wait : TIMER;   // Wait for glass process
   tmON_AuxFunction1 : TIMER;   // Timer auxiliary function 1
   tmON_AuxFunction2 : TIMER;   // Timer auxiliary function 2
   tmON_AuxFunction3 : TIMER;   // Timer auxiliary function 3
   tmON_AuxFunction4 : TIMER;   // Timer auxiliary function 4
   tmON_AuxFunction5 : TIMER;   // Timer auxiliary function 5
   tmON_AuxFunction6 : TIMER;   // Timer auxiliary function 6
   tmON_AuxFunction7 : TIMER;   // Timer auxiliary function 7
   tmON_AuxFunction8 : TIMER;   // Timer auxiliary function 8
   tmON_AuxFunction9 : TIMER;   // Timer auxiliary function 9
   tmOF_MCD_M1 : TIMER;
   tmOF_MCD_M2 : TIMER;
   tmOF_MCD_M3 : TIMER;
   tmOF_MCD_M4 : TIMER;
END_STRUCT
END_TYPE
